// TIA Portal project "EbAndon v4_00_038" (V15) (continued)
DEVICE "ET 200SP station_29"  ET 200SP-Station
   slot 0: "Rack_0"  Rack  6ES5 710-8MAx1
   slot 0: "cv04et200sp"  IM 155-6 PN ST  6ES7 155-6AU01-0BN0  V4.1
   slot 1: "DQ 8x24VDC/0.5A ST_1"  DQ 8x24VDC/0.5A ST  6ES7 132-6BF01-0BA0  V0.0
      slot 1: "DQ 8x24VDC/0.5A ST_1"  DQ 8x24VDC/0.5A ST
   slot 2: "DQ 8x24VDC/0.5A ST_2"  DQ 8x24VDC/0.5A ST  6ES7 132-6BF01-0BA0  V0.0
      slot 1: "DQ 8x24VDC/0.5A ST_2"  DQ 8x24VDC/0.5A ST
   slot 3: "DQ 8x24VDC/0.5A ST_3"  DQ 8x24VDC/0.5A ST  6ES7 132-6BF01-0BA0  V0.0
      slot 1: "DQ 8x24VDC/0.5A ST_3"  DQ 8x24VDC/0.5A ST
   slot 4: "Server module_1"  Server module  6ES7 193-6PA00-0AA0  V1.1
      slot 1: "Server module_1"  Server module
   slot 127: "BA 2xRJ45"  BA 2xRJ45  6ES7 193-6AR00-0AA0  V0.0
      slot 1: "Port_1"  6ES7 193-6AR00-0AA0  V0.0
      slot 2: "Port_2"  6ES7 193-6AR00-0AA0  V0.0
DEVICE "ET 200SP station_30"  ET 200SP-Station
   slot 0: "Rack_0"  Rack  6ES5 710-8MAx1
   slot 0: "pc01et200sp"  IM 155-6 PN ST  6ES7 155-6AU01-0BN0  V4.1
   slot 1: "DQ 8x24VDC/0.5A ST_1"  DQ 8x24VDC/0.5A ST  6ES7 132-6BF01-0BA0  V0.0
      slot 1: "DQ 8x24VDC/0.5A ST_1"  DQ 8x24VDC/0.5A ST
   slot 2: "DQ 8x24VDC/0.5A ST_2"  DQ 8x24VDC/0.5A ST  6ES7 132-6BF01-0BA0  V0.0
      slot 1: "DQ 8x24VDC/0.5A ST_2"  DQ 8x24VDC/0.5A ST
   slot 3: "DQ 8x24VDC/0.5A ST_3"  DQ 8x24VDC/0.5A ST  6ES7 132-6BF01-0BA0  V0.0
      slot 1: "DQ 8x24VDC/0.5A ST_3"  DQ 8x24VDC/0.5A ST
   slot 4: "Server module_1"  Server module  6ES7 193-6PA00-0AA0  V1.1
      slot 1: "Server module_1"  Server module
   slot 127: "BA 2xRJ45"  BA 2xRJ45  6ES7 193-6AR00-0AA0  V0.0
      slot 1: "Port_1"  6ES7 193-6AR00-0AA0  V0.0
      slot 2: "Port_2"  6ES7 193-6AR00-0AA0  V0.0
DEVICE "ET 200SP station_31"  ET 200SP-Station
   slot 0: "Rack_0"  Rack  6ES5 710-8MAx1
   slot 0: "pc02et200sp"  IM 155-6 PN ST  6ES7 155-6AU01-0BN0  V4.1
   slot 1: "DQ 8x24VDC/0.5A ST_1"  DQ 8x24VDC/0.5A ST  6ES7 132-6BF01-0BA0  V0.0
      slot 1: "DQ 8x24VDC/0.5A ST_1"  DQ 8x24VDC/0.5A ST
   slot 2: "DQ 8x24VDC/0.5A ST_2"  DQ 8x24VDC/0.5A ST  6ES7 132-6BF01-0BA0  V0.0
      slot 1: "DQ 8x24VDC/0.5A ST_2"  DQ 8x24VDC/0.5A ST
   slot 3: "DQ 8x24VDC/0.5A ST_3"  DQ 8x24VDC/0.5A ST  6ES7 132-6BF01-0BA0  V0.0
      slot 1: "DQ 8x24VDC/0.5A ST_3"  DQ 8x24VDC/0.5A ST
   slot 4: "Server module_1"  Server module  6ES7 193-6PA00-0AA0  V1.1
      slot 1: "Server module_1"  Server module
   slot 127: "BA 2xRJ45"  BA 2xRJ45  6ES7 193-6AR00-0AA0  V0.0
      slot 1: "Port_1"  6ES7 193-6AR00-0AA0  V0.0
      slot 2: "Port_2"  6ES7 193-6AR00-0AA0  V0.0
*)

// ===== PLC "PLC_1"  CPU 1517F-3 PN/DP =====

VAR_GLOBAL   // PLC tag table "Default tag table"
   "System_Byte" AT %MB1 : Byte;
   "FirstScan" AT %M1.0 : Bool;
   "DiagStatUpdt" AT %M1.1 : Bool;
   "AlwaysTRUE" AT %M1.2 : Bool;
   "AlwaysFALSE" AT %M1.3 : Bool;
   "Clock_Byte" AT %MB0 : Byte;
   "Clock_10Hz" AT %M0.0 : Bool;
   "Clock_5Hz" AT %M0.1 : Bool;
   "Clock_2.5Hz" AT %M0.2 : Bool;
   "Clock_2Hz" AT %M0.3 : Bool;
   "Clock_1.25Hz" AT %M0.4 : Bool;
   "Clock_1Hz" AT %M0.5 : Bool;
   "Clock_0.625Hz" AT %M0.6 : Bool;
   "Clock_0.5Hz" AT %M0.7 : Bool;
   "Temp Reset" AT %M2.0 : Bool;
   "clearPartData" AT %M100.0 : Bool;
   "setDefaultPresets" AT %M100.1 : Bool;
   "hardInitReq" AT %M100.2 : Bool;
   "dbg" AT %M500.0 : Bool;
   "dbgSetDefTimes" AT %M5000.0 : Bool;
   "Copy PN Codes Into Recipes" AT %M10.0 : Bool;
   "Load Default Recipes Into Stations" AT %M10.1 : Bool;
   "Load Default Wip Data" AT %M10.2 : Bool;
   "dbg_station_index" AT %MW502 : Int;
END_VAR

VAR_GLOBAL CONSTANT   // PLC tag table "Default tag table"
   "PARTS_PER_STATION" : Int := 7;
   "_SELECT_STATION_BUTTON_COUNT" : Int := 11;
   "NULL_TOKEN" : Int := -1;
   "WIP_POPUP_BUTTON_COUNT" : Int := 6;   // number of wip select buttons on wip select pop up screen
   "LINKED_LIST_LENGTH" : Int := 49;
   "SHOW" : Bool := TRUE;
   "HIDE" : Bool := FALSE;
   "BLANK" : WString := WSTRING#'';
END_VAR

VAR_GLOBAL   // PLC tag table "VOLVO 16 01"
   "VOLVO 16 01 IO" AT %QD1000 : DWord;
   "VOLVO 16 01 KP8 In" AT %ID0 : DWord;
   "VOLVO 16 01 KP8 Out" AT %QD0 : DWord;
END_VAR

VAR_GLOBAL   // PLC tag table "VOLVO 16 02"
   "VOLVO 16 02 IO" AT %QD1004 : DWord;
   "VOLVO 16 02 KP8 In" AT %ID4 : DWord;
   "VOLVO 16 02 KP8 Out" AT %QD4 : DWord;
END_VAR

VAR_GLOBAL   // PLC tag table "VOLVO 16 03"
   "VOLVO 16 03 IO" AT %QD1008 : DWord;
   "VOLVO 16 03 KP8 In" AT %ID8 : DWord;
   "VOLVO 16 03 KP8 Out" AT %QD8 : DWord;
END_VAR

VAR_GLOBAL   // PLC tag table "VOLVO 16 04"
   "VOLVO 16 04 IO" AT %QD1012 : DWord;
   "VOLVO 16 04 KP8 In" AT %ID12 : DWord;
   "VOLVO 16 04 KP8 Out" AT %QD12 : DWord;
END_VAR

VAR_GLOBAL   // PLC tag table "VOLVO 16 05"
   "VOLVO 16 05 IO" AT %QD1016 : DWord;
   "VOLVO 16 05 KP8 In" AT %ID16 : DWord;
   "VOLVO 16 05 KP8 Out" AT %QD16 : DWord;
END_VAR

VAR_GLOBAL   // PLC tag table "VOLVO 16 06"
   "VOLVO 16 06 IO" AT %QD1020 : DWord;
   "VOLVO 16 06 KP8 In" AT %ID20 : DWord;
   "VOLVO 16 06 KP8 Out" AT %QD20 : DWord;
END_VAR

VAR_GLOBAL   // PLC tag table "VOLVO 16 07"
   "VOLVO 16 07 IO" AT %QD1024 : DWord;
   "VOLVO 16 07 KP8 In" AT %ID24 : DWord;
   "VOLVO 16 07 KP8 Out" AT %QD24 : DWord;
END_VAR

VAR_GLOBAL   // PLC tag table "VOLVO 16 08"
   "VOLVO 16 08 IO" AT %QD1028 : DWord;
   "VOLVO 16 08 KP8 In" AT %ID28 : DWord;
   "VOLVO 16 08 KP8 Out" AT %QD28 : DWord;
END_VAR

VAR_GLOBAL   // PLC tag table "VOLVO 16 09"
   "VOLVO 16 09 IO" AT %QD1032 : DWord;
   "VOLVO 16 09 KP8 In" AT %ID32 : DWord;
   "VOLVO 16 09 KP8 Out" AT %QD32 : DWord;
END_VAR

VAR_GLOBAL   // PLC tag table "VOLVO 16 10"
   "VOLVO 16 10 IO" AT %QD1036 : DWord;
   "VOLVO 16 10 KP8 In" AT %ID36 : DWord;
   "VOLVO 16 10 KP8 Out" AT %QD36 : DWord;
END_VAR

VAR_GLOBAL   // PLC tag table "VOLVO 16 11"
   "VOLVO 16 11 IO" AT %QD1040 : DWord;
   "VOLVO 16 11 KP8 In" AT %ID40 : DWord;
   "VOLVO 16 11 KP8 Out" AT %QD40 : DWord;
END_VAR

VAR_GLOBAL   // PLC tag table "CHM 02"
   "CHM 02 KP8 In" AT %ID44 : DWord;
   "CHM 02 KP8 Out" AT %QD44 : DWord;
   "CHM 02 IO" AT %QD1044 : DWord;
END_VAR

VAR_GLOBAL   // PLC tag table "CHM 03"
   "CHM 03 IO" AT %QD1048 : DWord;
   "CHM 03 KP8 In" AT %ID48 : DWord;
   "CHM 03 KP8 Out" AT %QD48 : DWord;
END_VAR

VAR_GLOBAL   // PLC tag table "CHM 04"
   "CHM 04 IO" AT %QD1052 : DWord;
   "CHM 04 KP8 In" AT %ID52 : DWord;
   "CHM 04 KP8 Out" AT %QD52 : DWord;
END_VAR

VAR_GLOBAL   // PLC tag table "CHM 05"
   "CHM 05 IO" AT %QD1056 : DWord;
   "CHM 05 KP8 In" AT %ID56 : DWord;
   "CHM 05 KP8 Out" AT %QD56 : DWord;
END_VAR

VAR_GLOBAL   // PLC tag table "CDO 01"
   "CDO 01 IO" AT %QD1060 : DWord;
   "CDO 01 KP8 In" AT %ID60 : DWord;
   "CDO 01 KP8 Out" AT %QD60 : DWord;
END_VAR

VAR_GLOBAL   // PLC tag table "CDO 02"
   "CDO 02 IO" AT %QD1064 : DWord;
   "CDO 02 KP8 In" AT %ID64 : DWord;
   "CDO 02 KP8 Out" AT %QD64 : DWord;
END_VAR

VAR_GLOBAL   // PLC tag table "CDO 03"
   "CDO 03 IO" AT %QD1068 : DWord;
   "CDO 03 KP8 In" AT %ID68 : DWord;
   "CDO 03 KP8 Out" AT %QD68 : DWord;
END_VAR

VAR_GLOBAL   // PLC tag table "BFL 01"
   "BFL 01 IO" AT %QD1072 : DWord;
   "BFL 01 KP8 In" AT %ID72 : DWord;
   "BFL 01 KP8 Out" AT %QD72 : DWord;
   "Manual Operations Trigger" AT %M10.3 : Bool;
END_VAR

VAR_GLOBAL   // PLC tag table "BFL 02"
   "BFL 02 IO" AT %QD1076 : DWord;
   "BFL 02 KP8 In" AT %ID76 : DWord;
   "BFL 02 KP8 Out" AT %QD76 : DWord;
END_VAR

VAR_GLOBAL   // PLC tag table "BFL 03"
   "BFL 03 IO" AT %QD1080 : DWord;
   "BFL 03 KP8 In" AT %ID80 : DWord;
   "BFL 03 KP8 Out" AT %QD80 : DWord;
END_VAR

VAR_GLOBAL   // PLC tag table "LGS 01"
   "LGS 01 IO" AT %QD1084 : DWord;
   "LGS 01 KP8 In" AT %ID84 : DWord;
   "LGS 01 KP8 Out" AT %QD84 : DWord;
END_VAR

VAR_GLOBAL   // PLC tag table "LGS 02"
   "LGS 02 IO" AT %QD1088 : DWord;
   "LGS 02 KP8 In" AT %ID88 : DWord;
   "LGS 02 KP8 Out" AT %QD88 : DWord;
END_VAR

VAR_GLOBAL   // PLC tag table "CHM 01"
   "CHM 01 IO" AT %QD1092 : DWord;
   "CHM 01 KP8 In" AT %ID92 : DWord;
   "CHM 01 KP8 Out" AT %QD92 : DWord;
END_VAR

VAR_GLOBAL CONSTANT   // PLC tag table "Comm Diag"
   "pnioDeviceCount" : Int := 48;   // Upper limit of devices per HMI screen
   "USERDIAG_SLOTS_PER_SCREEN_UPPER_LIM" : Int := 31;   // Upper limit of slots per HMI screen
   "USERDIAG_SLOTS_PER_DEVICE_UPPER_LIM" : Int := 31;   // max number of modules per device
   "USERDIAG_DEVICES_PER_IO_SYSTEM_UPPER_LIM" : Int := 128;   // Upper limit of devices/slaves per IO-System/DP-Mastersystem
   "USERDIAG_SLOTS_PER_PLC_UPPER_LIM" : Int := 31;   // max number of local modules
   "USERDIAG_IO_SYSTEMS_UPPER_LIM" : Int := 1;   // Upper limit of IO-Systems/DP-Mastersystems
   "USERDIAG_IOSYSTEM_1" : Int := 1;   // Index for first IO-System/DP-Mastersystem
END_VAR

VAR_GLOBAL CONSTANT   // PLC tag table "Color Library"
   "BLACK_BLACK" : USInt := 0;
   "WHITE_BACKGROUND" : USInt := 1;
   "WHITE_FOREGROUND" : USInt := 2;
   "WHITE_FLASHING" : USInt := 3;
   "GRAY_BACKGROUND" : USInt := 4;
   "GRAY_FOREGROUND" : USInt := 5;
   "GRAY_FLASHING" : USInt := 6;
   "RED_LIGHT_BACKGROUND" : USInt := 7;
   "RED_LIGTH_FOREGROUND" : USInt := 8;
   "RED_LIGHT_FLASHING" : USInt := 9;
   "RED_BACKGROUND" : USInt := 10;
   "RED_FOREGROUND" : USInt := 11;
   "RED_FLASHING" : USInt := 12;
   "YELLOW_LIGHT_BACKGROUND" : USInt := 13;
   "YELLOW_LIGHT_FOREGROUND" : USInt := 14;
   "YELLOW_LIGHT_FLASHING" : USInt := 15;
   "YELLOW_BACKGROUND" : USInt := 16;
   "YELLOW_FOREGROUND" : USInt := 17;
   "YELLOW_FLASHING" : USInt := 18;
   "GREEN_LIGHT_BACKGROUND" : USInt := 19;
   "GREEN_LIGHT_FOREGROUND" : USInt := 20;
   "GREEN_LIGHT_FLASHING" : USInt := 21;
   "GREEN_BACKGROUND" : USInt := 22;
   "GREEN_FOREGROUND" : USInt := 23;
   "GREEN_FLASHING" : USInt := 24;
   "TEAL_LIGHT_BACKGROUND" : USInt := 25;
   "TEAL_LIGHT_FOREGROUND" : USInt := 26;
   "TEAL_LIGHT_FLASHING" : USInt := 27;
   "TEAL_BACKGROUND" : USInt := 28;
   "TEAL_FOREGROUND" : USInt := 29;
   "TEAL_FLASHING" : USInt := 30;
   "BLUE_LIGHT_BACKGROUND" : USInt := 31;
   "BLUE_LIGHT_FOREGROUND" : USInt := 32;
   "BLUE_LIGHT_FLASHING" : USInt := 33;
   "BLUE_BACKGROUND" : USInt := 34;
   "BLUE_FOREGROUND" : USInt := 35;
   "BLUE_FLASHING" : USInt := 36;
   "PURPLE_LIGHT_BACKGROUND" : USInt := 37;
   "PURPLE_LIGHT_FOREGROUND" : USInt := 38;   // foreground light purple
   "PURPLE_LIGHT_FLASHING" : USInt := 39;
   "PURPLE_DARK_BACKGROUND" : USInt := 40;
   "PURPLE_DARK_FOREGROUND" : USInt := 41;
   "PURPLE_FLASHING" : USInt := 42;
   "DISABLED" : USInt := 254;
   "INVISIBLE" : USInt := 255;
   "LBlDRd" : USInt := 43;
   "DRdLBl" : USInt := 44;
   "LBlDRdFl" : USInt := 45;
   "DBlDRd" : USInt := 46;
   "DRdDBl" : USInt := 47;
   "DBlDRdFl" : USInt := 48;
END_VAR

VAR_GLOBAL CONSTANT   // PLC tag table "Station Meta Data"
   "BUTTON_COUNT" : Int := 7;   // one less than actual button count
   "STATION_COUNT" : Int := 38;   // one less than actual station count
   "DEFAULT_TOTAL" : Real := 1800.0;
   "DEFAULT_CRITICAL" : Real := 300.0;
   "WIP_COUNT" : Int := 49;   // one less than actual wip count
   "MEDIUM_STRING_LENGTH" : Int := 40;
   "SHORT_STRING_LENGTH" : Int := 20;
   "LONG_STRING_LENGTH" : Int := 100;
   "PART_NUMBER_LIBRARY_COUNT" : Int := 999;   // one less than actual pn capacity
   "KP8_STATION_COUNT" : Int := 33;
   "HMI_STATION_COUNT" : Int := 4;   // number of stations using basic panel instead of kp8 (-1 for array)
END_VAR

VAR_GLOBAL   // PLC tag table "Simulation"
   "simMode" AT %M100.3 : Bool;
END_VAR

VAR_GLOBAL CONSTANT   // PLC tag table "Simulation"
   "simKP8Count" : Int := 11;
END_VAR

VAR_GLOBAL CONSTANT   // PLC tag table "Station IDs"
   "VOLVO 16 01" : Int := 0;
   "VOLVO 16 02" : Int := 1;
   "VOLVO 16 03" : Int := 2;
   "VOLVO 16 04" : Int := 3;
   "VOLVO 16 05" : Int := 4;
   "VOLVO 16 06" : Int := 5;
   "VOLVO 16 07" : Int := 6;
   "VOLVO 16 08" : Int := 7;
   "VOLVO 16 09" : Int := 8;
   "VOLVO 16 10" : Int := 9;
   "VOLVO 16 11" : Int := 10;
   "CHM 01" : Int := 11;
   "CHM 02" : Int := 12;
   "CHM 03" : Int := 13;
   "CHM 04" : Int := 14;
   "CHM 05" : Int := 15;
   "CDO 01" : Int := 16;
   "CDO 02" : Int := 17;
   "CDO 03" : Int := 18;
   "BFL 01" : Int := 19;
   "BFL 02" : Int := 20;
   "BFL 03" : Int := 21;
   "LGS 01" : Int := 22;
   "LGS 02" : Int := 23;
   "LGS 03" : Int := 24;
   "CV 01" : Int := 25;
   "CV 02" : Int := 26;
   "CV 03" : Int := 27;
   "CV 04" : Int := 28;
   "PC 01" : Int := 29;
   "PC 02" : Int := 30;
END_VAR

VAR_GLOBAL CONSTANT   // PLC tag table "LED Sign"
   "ledRowCount" : Int := 11;
END_VAR

VAR_GLOBAL CONSTANT   // PLC tag table "HMI Part Request Screen"
   "PART_REQUEST_ROW_COUNT_WAREHOUSE_HMI" : Int := 10;   // number of rows displayed on hmi
END_VAR

VAR_GLOBAL CONSTANT   // PLC tag table "HMI Settings Screen"
   "stngsScrnSlctdStns" : Int := 11;   // labels for settings screen
END_VAR

VAR_GLOBAL CONSTANT   // PLC tag table "Part Request Data Base"
   "partReqDataRowCount" : Int := 199;   // number of rows in part request table
END_VAR

VAR_GLOBAL CONSTANT   // PLC tag table "HMI Station"
   "wipSelScrnObjCnt" : Int := 29;   // number of buttons on menu select screen (short and long rows use different data, -1 for array)
   "partSelScrnObjCnt" : Int := 7;   // number of buttons on part select screen (-1 for array)
   "tmpltScrnObjCnt" : Int := 1;   // number of button on the template (-1 for array)
   "WIP_SELECT_BUTTON_COUNT" : Int := 5;   // button count for wip selection screen on hmi stations, -1 for array
END_VAR

VAR_GLOBAL   // PLC tag table "LGS 03"
   "LGS 03 IO" AT %QD1096 : DWord;
   "LGS 03 KP8 In" AT %ID96 : DWord;
   "LGS 03 KP8 Out" AT %QD96 : DWord;
END_VAR

VAR_GLOBAL   // PLC tag table "CV 01"
   "CV 01 IO" AT %QD1100 : DWord;
   "CV 01 KP8 In" AT %ID100 : DWord;
   "CV 01 KP8 Out" AT %QD100 : DWord;
END_VAR

VAR_GLOBAL   // PLC tag table "CV 02"
   "CV 02 IO" AT %QD1104 : DWord;
   "CV 02 KP8 In" AT %ID104 : DWord;
   "CV 02 KP8 Out" AT %QD104 : DWord;
END_VAR

VAR_GLOBAL   // PLC tag table "CV 03"
   "CV 03 IO" AT %QD1108 : DWord;
   "CV 03 KP8 In" AT %ID108 : DWord;
   "CV 03 KP8 Out" AT %QD108 : DWord;
END_VAR

VAR_GLOBAL   // PLC tag table "CV 04"
   "CV 04 IO" AT %QD1112 : DWord;
   "CV 04 KP8 In" AT %ID112 : DWord;
   "CV 04 KP8 Out" AT %QD112 : DWord;
END_VAR

VAR_GLOBAL   // PLC tag table "PC 01"
   "PC 01 IO" AT %QD1116 : DWord;
   "PC 01 KP8 In" AT %ID116 : DWord;
   "PC 01 KP8 Out" AT %QD116 : DWord;
END_VAR

VAR_GLOBAL   // PLC tag table "PC 02"
   "PC 02 IO" AT %QD1120 : DWord;
   "PC 02 KP8 In" AT %ID120 : DWord;
   "PC 02 KP8 Out" AT %QD120 : DWord;
END_VAR

VAR_GLOBAL CONSTANT   // PLC tag table "States"
   "requested" : Int := 10;
   "ordered" : Int := 20;
   "requestedCrit" : Int := 11;
   "requestedExp" : Int := 12;
   "acknowledged" : Int := 30;
   "reset" : Int := 99;
   "idle" : Int := 01;
   "orderedCrit" : Int := 21;
   "acknowledgedCrit" : Int := 31;
   "orderedExp" : Int := 22;
   "acknowledgedExp" : Int := 32;
END_VAR

VAR_GLOBAL CONSTANT   // PLC tag table "Timers"
   "DEFAULT_CRITICAL_TIME" : Real := 5.0;
   "DEFAULT_TOTAL_TIME" : Real := 10.0;
END_VAR

TYPE "Part Call Screen"
   STRUCT
      row : Array[0.."PART_REQUEST_ROW_COUNT_WAREHOUSE_HMI"] of "Table Row";
   END_STRUCT;
END_TYPE

TYPE "Barcode.UDT"
   STRUCT
      acknowledged : Bool;
      animate_acknowledged : Bool;
      animate_ordered : Bool;
      animate_cancel : Bool;
      address : DInt;
      barcode : String;
      color_acknowledged : UInt;
      color_ordered : UInt;
      color_cancel : UInt;
      ordered : Bool;
      part_number : WString[40];
   END_STRUCT;
END_TYPE

TYPE "Table Row"
   STRUCT
      address : DInt := -1;
      ordered : Bool;
      pbSelection : Struct
         actuate : Bool;
         animate : USInt;
      END_STRUCT;
      rtBackground : Struct
         animate : USInt;
      END_STRUCT;
      tfDropZone : Struct
         animate : USInt;
         value : WString[20];
      END_STRUCT;
      tfLine : Struct
         animate : USInt;
         value : WString[20];
      END_STRUCT;
      tfPartNumber : Struct
         animateDL : USInt;
         animateSL : USInt;
         value : WString[40];
      END_STRUCT;
      tfTime : Struct
         animate : USInt;
         value : WString[20];
      END_STRUCT;
   END_STRUCT;
END_TYPE

TYPE "Part Request Data"
   STRUCT
      row : Array[0.."partReqDataRowCount"] of DInt;
   END_STRUCT;
END_TYPE

TYPE "Settings"
   STRUCT
      selectStation : "Push Button Data";
      selectWip : "Push Button Data";
      selectButton : "Push Button Data";
      line : "IO Field Data: Label with Data";
      dropzone : "IO Field Data: Label with Data";
      total : "IO Field Data: Label with Data";
      critical : "IO Field Data: Label with Data";
      partNumber : "Part_Number_Double.UDT";
      assign : "Push Button Data";
      stationRows : Array[0..2] of "Settings Station Row Data";
      stnTableNavBar : "Nav Bar Data";
   END_STRUCT;
   // selectStation.animate := 1;
END_TYPE

TYPE "Push Button Data"
   STRUCT
      actuate : Bool;
      animate : USInt;
      enable : Bool;
      label : WString[80];
      listSelect : UInt;
      visible : Bool;
   END_STRUCT;
END_TYPE

TYPE "LED Sign Data"
   STRUCT
      row : Array[0.."ledRowCount"] of "Table Row";
   END_STRUCT;
END_TYPE

TYPE "Nav Bar Data: HMI"
   STRUCT
      top_actuate : Bool;
      top_animate : USInt;
      top_enable : Bool;
      top_label : WString;
      top_list_select : UInt;
      top_visible : Bool;
      page_up_actuate : Bool;
      page_up_animate : USInt;
      page_up_enable : Bool;
      page_up_label : WString;
      page_up_list_select : UInt;
      page_up_visible : Bool;
      line_up_actuate : Bool;
      line_up_animate : USInt;
      line_up_enable : Bool;
      line_up_label : WString;
      line_up_list_select : UInt;
      line_up_visible : Bool;
      line_down_actuate : Bool;
      line_down_animate : USInt;
      line_down_enable : Bool;
      line_down_label : WString;
      line_down_list_select : UInt;
      line_down_visible : Bool;
      page_down_actuate : Bool;
      page_down_animate : USInt;
      page_down_enable : Bool;
      page_down_label : WString;
      page_down_list_select : UInt;
      page_down_visible : Bool;
      bottom_actuate : Bool;
      bottom_animate : USInt;
      bottom_enable : Bool;
      bottom_label : WString;
      bottom_list_select : UInt;
      bottom_visible : Bool;
   END_STRUCT;
END_TYPE

TYPE "Pop Ups"
   STRUCT
      select_buttons : "Select Button";
      select_stations : "Select Station";
      select_WIPs : "Select WIP";
   END_STRUCT;
END_TYPE

TYPE "IO Field Data: Label with Data"
   STRUCT
      animate : USInt;
      enable : Bool;
      input_finished : Bool;
      value : WString[40];
      visible : Bool;
   END_STRUCT;
END_TYPE

TYPE "Selectable Station States"
   STRUCT
      all : Bool;
      non_hmi : Bool;
      hmi : Bool;
   END_STRUCT;
END_TYPE

TYPE "Selectable Stations"
   STRUCT
      count : Int;
      stns : Array[0.."STATION_COUNT"] of Int;
   END_STRUCT;
END_TYPE

TYPE "Nav Bar Data: PLC"
   STRUCT
      top : "Push Button Data";
      pageUp : "Push Button Data";
      lineUp : "Push Button Data";
      lineDown : "Push Button Data";
      pageDown : "Push Button Data";
      bottom : "Push Button Data";
   END_STRUCT;
END_TYPE

TYPE "Simulated Stations"
   STRUCT
      down : "Push Button Data";
      firstStn : Int;
      me : Array[0.."simKP8Count"] of "Station: Sim Data";
      up : "Push Button Data";
   END_STRUCT;
END_TYPE

TYPE "Runtime Data"
   STRUCT
      asReal : Real;
      elapsed : LReal;
      mem : LReal;
   END_STRUCT;
END_TYPE

TYPE "Recipe: Wip Text Library"
   STRUCT
      code : Array[0..99] of WString["SHORT_STRING_LENGTH"];
      txt : Array[0..99] of WString["LONG_STRING_LENGTH"];
   END_STRUCT;
END_TYPE

TYPE "Recipe: HMI Stations Saved Wips"
   STRUCT
      stn : Array[0.."HMI_STATION_COUNT"] of "WIP: Station";
   END_STRUCT;
END_TYPE

TYPE "Network Health Screen"
   STRUCT
      et200spPopUp : "Station: ET200SP Comm Debug Data";
      kp8PopUp : "Station: KP8 Comm Debug Data";
      pnioDevices : Array[1.."pnioDeviceCount"] of "Push Button Data";
      selectedDevice : Int;
   END_STRUCT;
END_TYPE

TYPE "ET200SP: IM Data"
   STRUCT
      bg : USInt;
      error : USInt;
      lnk01 : USInt;
      lnk02 : USInt;
      maint : USInt;
      pwr : USInt;
      run : USInt;
   END_STRUCT;
END_TYPE

TYPE "ET200SP: DQ Data"
   STRUCT
      bg : USInt;
      bgTem : USInt;
      diag : USInt;
      pwr : USInt;
      x0 : USInt;
      x1 : USInt;
      x2 : USInt;
      x3 : USInt;
      x4 : USInt;
      x5 : USInt;
      x6 : USInt;
      x7 : USInt;
   END_STRUCT;
END_TYPE

TYPE "ET200SP: Server Module Data"
   STRUCT
      bg : USInt;
   END_STRUCT;
END_TYPE

TYPE "Settings Station Row Data"
   STRUCT
      line : "Cell Data";
      dropzone : "Cell Data";
      wip : "Cell Data";
      btnRows : Array[0..7] of "Settings Station Row Button Row Data";
   END_STRUCT;
END_TYPE

TYPE "Selected Stations"
   STRUCT
      count : Int;
      stns : Array[0.."STATION_COUNT"] of Bool;
   END_STRUCT;
END_TYPE

TYPE "Cell Data"
   STRUCT
      animate : Int;
      data : WString [58];
      visibility : Bool;
   END_STRUCT;
END_TYPE

TYPE "Settings Station Row Button Row Data"
   STRUCT
      button : "Cell Data";
      total : "Cell Data";
      critical : "Cell Data";
      singlePN : "Cell Data";
      doublePN : "Cell Data";
   END_STRUCT;
END_TYPE

TYPE "Select Button"
   STRUCT
      close_screen : "Push Button Data";
      buttons : Array[0..7] of "Push Button Data";
   END_STRUCT;
END_TYPE

TYPE "Select Station"
   STRUCT
      close_screen : "Push Button Data";
      nav_bar : "Nav Bar Data";
      stn_select_btns : Array[0.."_SELECT_STATION_BUTTON_COUNT"] of "Push Button Data";
   END_STRUCT;
END_TYPE

TYPE "Select WIP"
   STRUCT
      close_screen : "Push Button Data";
      nav_bar : "Nav Bar Data";
      select_wip_buttons : Array[0.."WIP_POPUP_BUTTON_COUNT"] of "Push Button Data";
   END_STRUCT;
END_TYPE

TYPE "WIP: Station"
   STRUCT
      pStn : Int;
      wip : Array[0.."WIP_COUNT"] of "Station: Wip: Wip Module";
   END_STRUCT;
END_TYPE

TYPE "Selectable Wips"
   STRUCT
      count : Int;
      wips : Array[0.."WIP_COUNT"] of DInt;
   END_STRUCT;
END_TYPE

TYPE "Recipe: PN Text Library"
VERSION : 0.1
   STRUCT
      pnText : Array[0.."PART_NUMBER_LIBRARY_COUNT"] of WString["SHORT_STRING_LENGTH"];
   END_STRUCT;
   // pnText[0] := WSTRING#'//';
   // pnText[1] := WSTRING#'//';
   // pnText[2] := WSTRING#'//';
   // pnText[3] := WSTRING#'//';
   // pnText[4] := WSTRING#'//';
   // pnText[5] := WSTRING#'//';
   // pnText[6] := WSTRING#'//';
   // pnText[7] := WSTRING#'//';
   // pnText[8] := WSTRING#'//';
   // pnText[9] := WSTRING#'//';
   // pnText[10] := WSTRING#'//';
   // pnText[11] := WSTRING#'//';
   // pnText[12] := WSTRING#'//';
   // pnText[13] := WSTRING#'//';
   // pnText[14] := WSTRING#'//';
   // pnText[15] := WSTRING#'//';
   // pnText[16] := WSTRING#'//';
   // pnText[17] := WSTRING#'//';
   // pnText[18] := WSTRING#'//';
   // pnText[19] := WSTRING#'//';
   // pnText[20] := WSTRING#'//';
   // pnText[21] := WSTRING#'//';
   // pnText[22] := WSTRING#'//';
   // pnText[23] := WSTRING#'//';
   // pnText[24] := WSTRING#'//';
   // pnText[25] := WSTRING#'//';
   // pnText[26] := WSTRING#'//';
   // pnText[27] := WSTRING#'//';
   // pnText[28] := WSTRING#'//';
   // pnText[29] := WSTRING#'//';
   // pnText[30] := WSTRING#'//';
   // pnText[31] := WSTRING#'//';
   // pnText[32] := WSTRING#'//';
   // pnText[33] := WSTRING#'//';
   // pnText[34] := WSTRING#'//';
   // pnText[35] := WSTRING#'//';
   // pnText[36] := WSTRING#'//';
   // pnText[37] := WSTRING#'//';
   // pnText[38] := WSTRING#'//';
   // pnText[39] := WSTRING#'//';
   // pnText[40] := WSTRING#'//';
   // pnText[41] := WSTRING#'//';
   // pnText[42] := WSTRING#'//';
   // pnText[43] := WSTRING#'//';
   // pnText[44] := WSTRING#'//';
   // pnText[45] := WSTRING#'//';
   // pnText[46] := WSTRING#'//';
   // pnText[47] := WSTRING#'//';
   // pnText[48] := WSTRING#'//';
   // pnText[49] := WSTRING#'//';
   // pnText[50] := WSTRING#'//';
   // pnText[51] := WSTRING#'//';
   // pnText[52] := WSTRING#'//';
   // pnText[53] := WSTRING#'//';
   // pnText[54] := WSTRING#'//';
   // pnText[55] := WSTRING#'//';
   // pnText[56] := WSTRING#'//';
   // pnText[57] := WSTRING#'//';
   // pnText[58] := WSTRING#'//';
   // pnText[59] := WSTRING#'//';
   // pnText[60] := WSTRING#'//';
   // pnText[61] := WSTRING#'//';
   // pnText[62] := WSTRING#'//';
   // pnText[63] := WSTRING#'//';
   // pnText[64] := WSTRING#'//';
   // pnText[65] := WSTRING#'//';
   // pnText[66] := WSTRING#'//';
   // pnText[67] := WSTRING#'//';
   // pnText[68] := WSTRING#'//';
   // pnText[69] := WSTRING#'//';
   // pnText[70] := WSTRING#'//';
   // pnText[71] := WSTRING#'//';
   // pnText[72] := WSTRING#'//';
   // pnText[73] := WSTRING#'//';
   // pnText[74] := WSTRING#'//';
   // pnText[75] := WSTRING#'//';
   // pnText[76] := WSTRING#'//';
   // pnText[77] := WSTRING#'//';
   // pnText[78] := WSTRING#'//';
   // pnText[79] := WSTRING#'//';
   // pnText[80] := WSTRING#'//';
   // pnText[81] := WSTRING#'//';
   // pnText[82] := WSTRING#'//';
   // pnText[83] := WSTRING#'//';
   // pnText[84] := WSTRING#'//';
   // pnText[85] := WSTRING#'//';
   // pnText[86] := WSTRING#'//';
   // pnText[87] := WSTRING#'//';
   // pnText[88] := WSTRING#'//';
   // pnText[89] := WSTRING#'//';
   // pnText[90] := WSTRING#'//';
   // pnText[91] := WSTRING#'//';
   // pnText[92] := WSTRING#'//';
   // pnText[93] := WSTRING#'//';
   // pnText[94] := WSTRING#'//';
   // pnText[95] := WSTRING#'//';
   // pnText[96] := WSTRING#'//';
   // pnText[97] := WSTRING#'//';
   // pnText[98] := WSTRING#'//';
   // pnText[99] := WSTRING#'//';
   // pnText[100] := WSTRING#'//';
   // pnText[101] := WSTRING#'//';
   // pnText[102] := WSTRING#'//';
   // pnText[103] := WSTRING#'//';
   // pnText[104] := WSTRING#'//';
   // pnText[105] := WSTRING#'//';
   // pnText[106] := WSTRING#'//';
   // pnText[107] := WSTRING#'//';
   // pnText[108] := WSTRING#'//';
   // pnText[109] := WSTRING#'//';
   // pnText[110] := WSTRING#'//';
   // pnText[111] := WSTRING#'//';
   // pnText[112] := WSTRING#'//';
   // pnText[113] := WSTRING#'//';
   // pnText[114] := WSTRING#'//';
   // pnText[115] := WSTRING#'//';
   // pnText[116] := WSTRING#'//';
   // pnText[117] := WSTRING#'//';
   // pnText[118] := WSTRING#'//';
   // pnText[119] := WSTRING#'//';
   // pnText[120] := WSTRING#'//';
   // pnText[121] := WSTRING#'//';
   // pnText[122] := WSTRING#'//';
   // pnText[123] := WSTRING#'//';
   // pnText[124] := WSTRING#'//';
   // pnText[125] := WSTRING#'//';
   // pnText[126] := WSTRING#'//';
   // pnText[127] := WSTRING#'//';
   // pnText[128] := WSTRING#'//';
   // pnText[129] := WSTRING#'//';
   // pnText[130] := WSTRING#'//';
   // pnText[131] := WSTRING#'//';
   // pnText[132] := WSTRING#'//';
   // pnText[133] := WSTRING#'//';
   // pnText[134] := WSTRING#'//';
   // pnText[135] := WSTRING#'//';
   // pnText[136] := WSTRING#'//';
   // pnText[137] := WSTRING#'//';
   // pnText[138] := WSTRING#'//';
   // pnText[139] := WSTRING#'//';
   // pnText[140] := WSTRING#'//';
   // pnText[141] := WSTRING#'//';
   // pnText[142] := WSTRING#'//';
   // pnText[143] := WSTRING#'//';
   // pnText[144] := WSTRING#'//';
   // pnText[145] := WSTRING#'//';
   // pnText[146] := WSTRING#'//';
   // pnText[147] := WSTRING#'//';
   // pnText[148] := WSTRING#'//';
   // pnText[149] := WSTRING#'//';
   // pnText[150] := WSTRING#'//';
   // pnText[151] := WSTRING#'//';
   // pnText[152] := WSTRING#'//';
   // pnText[153] := WSTRING#'//';
   // pnText[154] := WSTRING#'//';
   // pnText[155] := WSTRING#'//';
   // pnText[156] := WSTRING#'//';
   // pnText[157] := WSTRING#'//';
   // pnText[158] := WSTRING#'//';
   // pnText[159] := WSTRING#'//';
   // pnText[160] := WSTRING#'//';
   // pnText[161] := WSTRING#'//';
   // pnText[162] := WSTRING#'//';
   // pnText[163] := WSTRING#'//';
   // pnText[164] := WSTRING#'//';
   // pnText[165] := WSTRING#'//';
   // pnText[166] := WSTRING#'//';
   // pnText[167] := WSTRING#'//';
   // pnText[168] := WSTRING#'//';
   // pnText[169] := WSTRING#'//';
   // pnText[170] := WSTRING#'//';
   // pnText[171] := WSTRING#'//';
   // pnText[172] := WSTRING#'//';
   // pnText[173] := WSTRING#'//';
   // pnText[174] := WSTRING#'//';
   // pnText[175] := WSTRING#'//';
   // pnText[176] := WSTRING#'//';
   // pnText[177] := WSTRING#'//';
   // pnText[178] := WSTRING#'//';
   // pnText[179] := WSTRING#'//';
   // pnText[180] := WSTRING#'//';
   // pnText[181] := WSTRING#'//';
   // pnText[182] := WSTRING#'//';
   // pnText[183] := WSTRING#'//';
   // pnText[184] := WSTRING#'//';
   // pnText[185] := WSTRING#'//';
   // pnText[186] := WSTRING#'//';
   // pnText[187] := WSTRING#'//';
   // pnText[188] := WSTRING#'//';
   // pnText[189] := WSTRING#'//';
   // pnText[190] := WSTRING#'//';
   // pnText[191] := WSTRING#'//';
   // pnText[192] := WSTRING#'//';
   // pnText[193] := WSTRING#'//';
   // pnText[194] := WSTRING#'//';
   // pnText[195] := WSTRING#'//';
   // pnText[196] := WSTRING#'//';
   // pnText[197] := WSTRING#'//';
   // pnText[198] := WSTRING#'//';
   // pnText[199] := WSTRING#'//';
   // pnText[200] := WSTRING#'//';
   // pnText[201] := WSTRING#'//';
   // pnText[202] := WSTRING#'//';
   // pnText[203] := WSTRING#'//';
   // pnText[204] := WSTRING#'//';
   // pnText[205] := WSTRING#'//';
   // pnText[206] := WSTRING#'//';
   // pnText[207] := WSTRING#'//';
   // pnText[208] := WSTRING#'//';
   // pnText[209] := WSTRING#'//';
   // pnText[210] := WSTRING#'//';
   // pnText[211] := WSTRING#'//';
   // pnText[212] := WSTRING#'//';
   // pnText[213] := WSTRING#'//';
   // pnText[214] := WSTRING#'//';
   // pnText[215] := WSTRING#'//';
   // pnText[216] := WSTRING#'//';
   // pnText[217] := WSTRING#'//';
   // pnText[218] := WSTRING#'//';
   // pnText[219] := WSTRING#'//';
   // pnText[220] := WSTRING#'//';
   // pnText[221] := WSTRING#'//';
   // pnText[222] := WSTRING#'//';
   // pnText[223] := WSTRING#'//';
   // pnText[224] := WSTRING#'//';
   // pnText[225] := WSTRING#'//';
   // pnText[226] := WSTRING#'//';
   // pnText[227] := WSTRING#'//';
   // pnText[228] := WSTRING#'//';
   // pnText[229] := WSTRING#'//';
   // pnText[230] := WSTRING#'//';
   // pnText[231] := WSTRING#'//';
   // pnText[232] := WSTRING#'//';
   // pnText[233] := WSTRING#'//';
   // pnText[234] := WSTRING#'//';
   // pnText[235] := WSTRING#'//';
   // pnText[236] := WSTRING#'//';
   // pnText[237] := WSTRING#'//';
   // pnText[238] := WSTRING#'//';